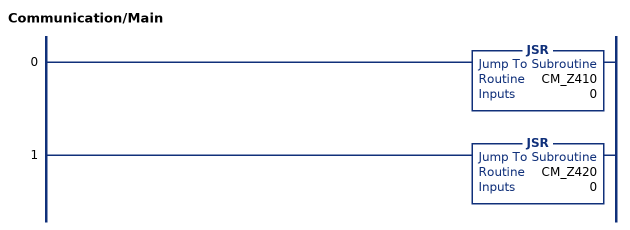
   0: JSR(CM_Z410,0);
   1: JSR(CM_Z420,0);
END_ROUTINE
END_PROGRAM

PROGRAM Initialize   (* main routine Main *)
VAR
   CapsConveyor_INIT : UDT_CapsConveyor_ZC[10]; {access None}
   Conveyor_INIT : UDT_StandConv[29]; {access None}
   M302SpeedUp_INIT : MAC_SpeedUp := (tmON_TimeControlSnap[0].PRE := 30000, tmON_TimeControlSnap[1].PRE := 30000); {constant, access None}
   M307ASpeedUp_INIT : MAC_SpeedUp := (tmON_TimeControlSnap[0].PRE := 30000, tmON_TimeControlSnap[1].PRE := 30000); {constant, access None}
   M30xTrimDeck_INIT : MAC_TrimmingDeck; {constant}
   M30xTrimWheels_INIT : MAC_TrimmingWheels[4]; {constant, access None}
        [1]   // M303 DW
        [2]   // M304 UP
        [3]   // M304 DW
        [0]   // M303 UP
   M310Popup_INIT : MAC_Popup_ZC[2]; {constant, access None}
        [0].PH_x.24   // Unload to stacker
        [0].PH_x.0   // Lift
        [0].PH_x.27   // End load to stacker
        [0].PH_x.16   // Squaring
        [0].PH_x.11   // Unload on side leg to opposite operator side
        [0].PH_x.15   // End unload to side leg
        [0].PH_x.19   // Positiong after squaring
        [0].PH_x.28   // Load from stacker
        [0].PH_x.3   // End lift
        [0].PH_x.31   // End load from stacker
        [0].PH_x.4   // Descent
        [0].PH_x.7   // End descent
        [0].PH_x.8   // Unload on side leg to operator side
        [1].PH_x.0   // Lift
        [1].PH_x.11   // Unload on side leg to opposite operator side
        [1].PH_x.15   // End unload to side leg
        [1].PH_x.16   // Squaring
        [1].PH_x.19   // Positiong after squaring
        [1].PH_x.24   // Unload to stacker
        [1].PH_x.27   // End load to stacker
        [1].PH_x.28   // Load from stacker
        [1].PH_x.3   // End lift
        [1].PH_x.31   // End load from stacker
        [1].PH_x.4   // Descent
        [1].PH_x.7   // End descent
        [1].PH_x.8   // Unload on side leg to operator side
   M315Popup_INIT : MAC_Popup_ZC[2]; {constant, access None}
        [0].PH_x.0   // Lift
        [0].PH_x.11   // Unload on side leg to opposite operator side
        [0].PH_x.15   // End unload to side leg
        [0].PH_x.16   // Squaring
        [0].PH_x.19   // Positiong after squaring
        [0].PH_x.24   // Unload to stacker
        [0].PH_x.27   // End load to stacker
        [0].PH_x.28   // Load from stacker
        [0].PH_x.3   // End lift
        [0].PH_x.31   // End load from stacker
        [0].PH_x.4   // Descent
        [0].PH_x.7   // End descent
        [0].PH_x.8   // Unload on side leg to operator side
        [1].PH_x.0   // Lift
        [1].PH_x.11   // Unload on side leg to opposite operator side
        [1].PH_x.15   // End unload to side leg
        [1].PH_x.16   // Squaring
        [1].PH_x.19   // Positiong after squaring
        [1].PH_x.24   // Unload to stacker
        [1].PH_x.27   // End load to stacker
        [1].PH_x.28   // Load from stacker
        [1].PH_x.3   // End lift
        [1].PH_x.31   // End load from stacker
        [1].PH_x.4   // Descent
        [1].PH_x.7   // End descent
        [1].PH_x.8   // Unload on side leg to operator side
   M350Popup_INIT : MAC_Popup_ZC; {access Read Only}
   Tracking_INIT : UDT_Tracking; {access None}
   Z301_INIT : MAC_Zone_ML := (tmON_ResetAlarm.PRE := 2000, tmON_24Vdc.PRE := 2000, tmON_400Vca.PRE := 2000, tmON_EmergencyOK.PRE := 2000, tmON_Cycle.PRE := 15000, tmON_ForceStop.PRE := 2000, tmON_AllowStopCleaning.PRE := 2000, tmON_CycleAcousticAlarm.PRE := 15000, tmON_ConveyorsNotOK.PRE := 2000, tmON_StopCycleForFaults.PRE := 2000, tmON_StopCycleForSaturation.PRE := 2000); {constant, access None}
END_VAR

ROUTINE Main   (* ladder *)
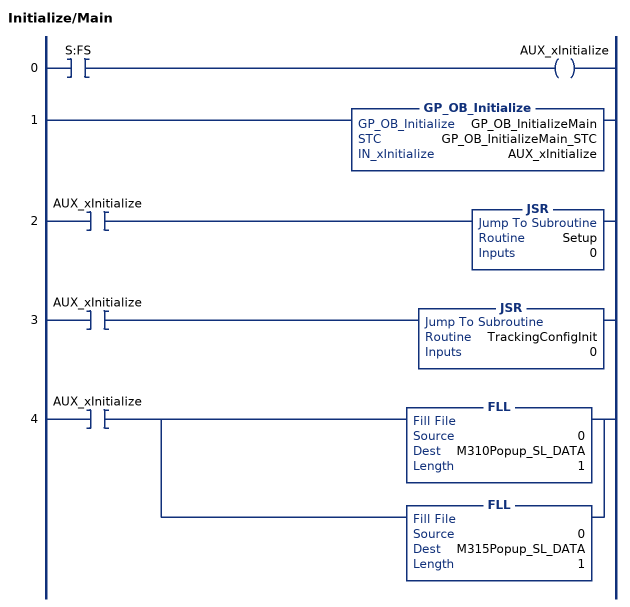
   0: XIC(S:FS)OTE(AUX_xInitialize);
   1: GP_OB_Initialize(GP_OB_InitializeMain,GP_OB_InitializeMain_STC,AUX_xInitialize);
   2: XIC(AUX_xInitialize)JSR(Setup,0);
   3: XIC(AUX_xInitialize)JSR(TrackingConfigInit,0);
   4: XIC(AUX_xInitialize)[FLL(0,M310Popup_SL_DATA,1) ,FLL(0,M315Popup_SL_DATA,1) ];
END_ROUTINE

ROUTINE Setup   (* structured text *)
   //Upload initialize parameters
   //Main line
   (*COP(Z301,Z301_INIT,1);
   COP(Z302,Z302_INIT,1);
   COP(Z303,Z303_INIT,1);
   COP(M301SpeedUp,M301SpeedUp_INIT,1);
   COP(M313SpeedUp,M313SpeedUp_INIT,1);
   COP(M31xConveyor[0],M31xConveyor_INIT[0],CONST_tPlant.dZ1ConveyorNumber);
   COP(M32xConveyor[0],M32xConveyor_INIT[0],CONST_tPlant.dZ2ConveyorNumber);
   COP(M33xConveyor[0],M33xConveyor_INIT[0],CONST_tPlant.dZ3ConveyorNumber);
   COP(M303TrimDeck,M303TrimDeck_INIT,1);
   COP(M303xTrimWheel[0],M303xTrimWheel_INIT[0],CONST_tPlant.dTrimWheelsNumber);
   COP(M311ASplitBar,M311ASplitBar_INIT,1);
   COP(M311BSeparatorRolls,M311BSeparatorRolls_INIT,1);
   COP(M385PowderMachine,M385_INIT,1);
   COP(M314AInputBreaker,M314AInputBreaker_INIT,1);
   COP(M320AInputBreaker,M320AInputBreaker_INIT,1);
   COP(M317Popup[0],M317Popup_INIT[0],2);
   COP(M325Popup[0],M325Popup_INIT[0],2);
   COP(M323Popup,M323Popup_INIT,1);
   COP(M327Popup,M327Popup_INIT,1);
   COP(M314BBreaker,M314BBreaker_INIT,1);
   COP(M320BBreaker,M320BBreaker_INIT,1);
   COP(M390Breaker,M390Breaker_INIT,1);*)
   
   //Download initialize parameters
   //Main line
   //COP(M31xConveyor_INIT[0],M31xConveyor[0],CONST_tPlant.dZ1ConveyorNumber);
   //COP(M32xConveyor_INIT[0],M32xConveyor[0],CONST_tPlant.dZ2ConveyorNumber);
   //COP(M33xConveyor_INIT[0],M33xConveyor[0],CONST_tPlant.dZ3ConveyorNumber);
   COP(Conveyor_INIT[0],Z300_Conveyor[0],CONST_tPlant.dNumOfConveyors);
   FOR TMP_dIndexConv := 0 TO CONST_tPlant.dNumOfConveyors - 1 DO
   	FOR TMP_dIndexCapConv := 0 TO CONST_tPlant.dNumCapsConveyor - 1 DO
   		COP(AUX_tCapsConveyor_NULL,Z300_LineTracking.rgtTrkConv[TMP_dIndexConv].Cap[TMP_dIndexCapConv],1);
   	END_FOR;
   END_FOR;
   COP(Z301_INIT,Z301,1);
   Z301.ST_xSelAutoMode:=1;
   
   COP(M302SpeedUp_INIT,M302SpeedUp,1);
   COP(M307ASpeedUp_INIT,M307ASpeedUp,1);
   FOR TMP_dIndex := 0 TO CONST_tPlant.dTrimDeckNumber - 1 DO
   	COP(M30xTrimDeck_INIT,M30xTrimDeck[TMP_dIndex],1);
   END_FOR;
   FOR TMP_dIndex := 0 TO CONST_tPlant.dTrimWheelsNumber - 1 DO
   	COP(M30xTrimWheels_INIT[0],M30xTrimWheel[TMP_dIndex],1);
   END_FOR;
   
   COP(M350Popup_INIT,M350Popup,1);
   
   FOR TMP_dIndex := 0 TO 1 DO
   	COP(M310Popup_INIT[0],M310Popup[TMP_dIndex],1);
   	COP(M315Popup_INIT[0],M315Popup[TMP_dIndex],1);
   END_FOR;
   
   (*//Preset time on indexed machines
   //Load preset time on M31xConveyors
   FOR TMP_dPnt1:=0 TO CONST_tPlant.dZ1ConveyorNumber - 1 DO
   	M31xConveyor[TMP_dPnt1].tmON_Wait.PRE:=0;
   	M31xConveyor[TMP_dPnt1].tmON_SyncTimeout.PRE:=20000;
   	M31xConveyor[TMP_dPnt1].tmOF_SyncTimeout.PRE:=2000;
   	M31xConveyor[TMP_dPnt1].tmON_PhFilter.PRE:=200;
   	IF M31xConveyor[TMP_dPnt1].CONST_dMotorNumber > 0 THEN
   		TMP_d:=M31xConveyor[TMP_dPnt1].CONST_dMotorNumber;
   	ELSE
   		TMP_d:=1;
   	END_IF;
   	FOR TMP_dPnt2:=0 TO TMP_d - 1 DO
   		M31xConveyor[TMP_dPnt1].tmON_FeedbackTimeOut[TMP_dPnt2].PRE:=1500;
   		M31xConveyor[TMP_dPnt1].tmOF_DriveEnable[TMP_dPnt2].PRE:=20000;
   	END_FOR;
   END_FOR;
   
   //Load preset time on M32xConveyors
   FOR TMP_dPnt1:=0 TO CONST_tPlant.dZ2ConveyorNumber - 1 DO
   	M32xConveyor[TMP_dPnt1].tmON_Wait.PRE:=0;
   	M32xConveyor[TMP_dPnt1].tmON_SyncTimeout.PRE:=20000;
   	M32xConveyor[TMP_dPnt1].tmOF_SyncTimeout.PRE:=2000;
   	M32xConveyor[TMP_dPnt1].tmON_PhFilter.PRE:=200;
   	IF M32xConveyor[TMP_dPnt1].CONST_dMotorNumber > 0 THEN
   		TMP_d:=M32xConveyor[TMP_dPnt1].CONST_dMotorNumber;
   	ELSE
   		TMP_d:=1;
   	END_IF;
   	FOR TMP_dPnt2:=0 TO TMP_d - 1 DO
   		M32xConveyor[TMP_dPnt1].tmON_FeedbackTimeOut[TMP_dPnt2].PRE:=1500;
   		M32xConveyor[TMP_dPnt1].tmOF_DriveEnable[TMP_dPnt2].PRE:=20000;
   	END_FOR;
   END_FOR;
   
   //Load preset time on M33xConveyors
   FOR TMP_dPnt1:=0 TO CONST_tPlant.dZ2ConveyorNumber - 1 DO
   	M33xConveyor[TMP_dPnt1].tmON_Wait.PRE:=0;
   	M33xConveyor[TMP_dPnt1].tmON_SyncTimeout.PRE:=20000;
   	M33xConveyor[TMP_dPnt1].tmOF_SyncTimeout.PRE:=2000;
   	M33xConveyor[TMP_dPnt1].tmON_PhFilter.PRE:=200;
   	IF M33xConveyor[TMP_dPnt1].CONST_dMotorNumber > 0 THEN
   		TMP_d:=M33xConveyor[TMP_dPnt1].CONST_dMotorNumber;
   	ELSE
   		TMP_d:=1;
   	END_IF;
   	FOR TMP_dPnt2:=0 TO TMP_d - 1 DO
   		M33xConveyor[TMP_dPnt1].tmON_FeedbackTimeOut[TMP_dPnt2].PRE:=1500;
   		M33xConveyor[TMP_dPnt1].tmOF_DriveEnable[TMP_dPnt2].PRE:=20000;
   	END_FOR;
   END_FOR;*)
   
   //Load preset time on M30xTrimDeck
   FOR TMP_d :=0 TO CONST_tPlant.dTrimDeckNumber - 1 DO
   	M30xTrimDeck[TMP_d].tmON_EncPreset[0].PRE:=3000;
   	M30xTrimDeck[TMP_d].tmON_EncPreset[1].PRE:=3000;
   	M30xTrimDeck[TMP_d].tmON_CheckEncoderTimeOut[0].PRE:=1000;
   	M30xTrimDeck[TMP_d].tmON_CheckEncoderTimeOut[1].PRE:=1000;
   	M30xTrimDeck[TMP_d].tmON_FeedbackTimeOut[0].PRE:=2500;
   	M30xTrimDeck[TMP_d].tmON_FeedbackTimeOut[1].PRE:=2500;
   	M30xTrimDeck[TMP_d].tmOF_DriveEnable[0].PRE:=30000;
   	M30xTrimDeck[TMP_d].tmOF_DriveEnable[1].PRE:=30000;
   	M30xTrimDeck[TMP_d].tmOF_DelayOnChangeDirection[0].PRE:=500;
   	M30xTrimDeck[TMP_d].tmOF_DelayOnChangeDirection[1].PRE:=500;
   	M30xTrimDeck[TMP_d].tmOF_DelayOnChangeDirection[2].PRE:=500;
   	M30xTrimDeck[TMP_d].tmOF_DelayOnChangeDirection[3].PRE:=500;
   	M30xTrimDeck[TMP_d].tmON_Wait.PRE:=0;
   END_FOR;
   
   //Load preset time on M30xTrimWheels
   FOR TMP_d :=0 TO CONST_tPlant.dTrimWheelsNumber - 1 DO
   	M30xTrimWheel[TMP_d].tmON_TrimWheelTimeOut[0].PRE:=2500;
   	M30xTrimWheel[TMP_d].tmON_TrimWheelTimeOut[1].PRE:=2500;
   	M30xTrimWheel[TMP_d].tmON_Wait[0].PRE:=0;
   	M30xTrimWheel[TMP_d].tmON_Wait[1].PRE:=0;
   END_FOR;
   
   //Load preset time M317Popup
   M310Popup[0].tmON_LiftingTimeOut.PRE := 2000;
   M310Popup[0].tmON_LiftingFeedbackTimeOut.PRE := 1000;
   M310Popup[0].tmOF_WaitBothEndLift.PRE := 1500;
   M310Popup[0].tmON_ReentryPlate.PRE := 200;
   M310Popup[0].tmON_Positioning.PRE := 40;
   M310Popup[1].tmON_LiftingTimeOut.PRE := 2000;
   M310Popup[1].tmON_LiftingFeedbackTimeOut.PRE := 1000;
   M310Popup[1].tmOF_WaitBothEndLift.PRE := 1500;
   M310Popup[1].tmON_ReentryPlate.PRE := 200;
   M310Popup[1].tmON_Positioning.PRE := 40;
   
   //Load preset time M325Popup
   M315Popup[0].tmON_LiftingTimeOut.PRE := 2000;
   M315Popup[0].tmON_LiftingFeedbackTimeOut.PRE := 1000;
   M315Popup[0].tmOF_WaitBothEndLift.PRE := 1500;
   M315Popup[0].tmON_ReentryPlate.PRE := 200;
   M315Popup[0].tmON_Positioning.PRE := 40;
   M315Popup[1].tmON_LiftingTimeOut.PRE := 2000;
   M315Popup[1].tmON_LiftingFeedbackTimeOut.PRE := 1000;
   M315Popup[1].tmOF_WaitBothEndLift.PRE := 1500;
   M315Popup[1].tmON_ReentryPlate.PRE := 200;
   M315Popup[1].tmON_Positioning.PRE := 40;
   
END_ROUTINE

ROUTINE TrackingConfigInit   (* structured text *)
   
   Z300_dStartTrackingPosition := 0;
   Z300_LineTracking.rgtTrkConv[0].dStartPosition_cmm := Z300_dStartTrackingPosition;
   Z300_LineTracking.rgtTrkConv[0].dEndPosition_cmm := Z300_dStartTrackingPosition + Z300_Conveyor_Conf[0].dLengthConveyor_cmm;
   size(Z300_LineTracking.rgtTrkConv[0],0,TMP_dLineSize);
   FOR TMP_dIndexConv := 1 TO TMP_dLineSize - 1 DO
   	Z300_LineTracking.rgtTrkConv[TMP_dIndexConv].dStartPosition_cmm := Z300_LineTracking.rgtTrkConv[TMP_dIndexConv - 1].dEndPosition_cmm;
   	Z300_LineTracking.rgtTrkConv[TMP_dIndexConv].dEndPosition_cmm := Z300_LineTracking.rgtTrkConv[TMP_dIndexConv].dStartPosition_cmm + Z300_Conveyor_Conf[TMP_dIndexConv].dLengthConveyor_cmm;
   END_FOR;
   Z300_dEndTrackingPosition := Z300_LineTracking.rgtTrkConv[TMP_dLineSize - 1].dEndPosition_cmm;
   
END_ROUTINE
END_PROGRAM

PROGRAM MainProgram   (* main routine MainRoutine *)

ROUTINE _10_MCP_I   (* ladder *)
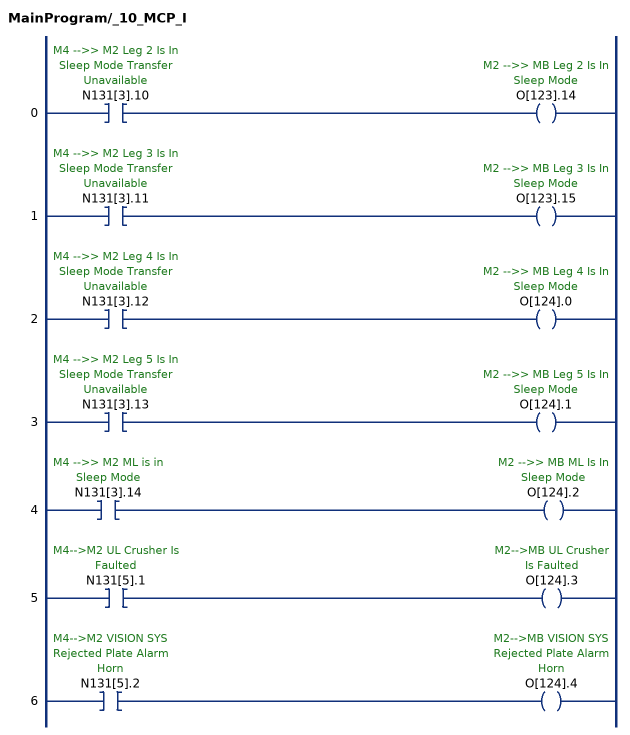
   0: XIC(N131[3].10)OTE(O[123].14);
   1: XIC(N131[3].11)OTE(O[123].15);
   2: XIC(N131[3].12)OTE(O[124].0);
   3: XIC(N131[3].13)OTE(O[124].1);
   4: XIC(N131[3].14)OTE(O[124].2);
   5: XIC(N131[5].1)OTE(O[124].3);
   6: XIC(N131[5].2)OTE(O[124].4);
END_ROUTINE

ROUTINE _12_MCP_K   (* ladder *)
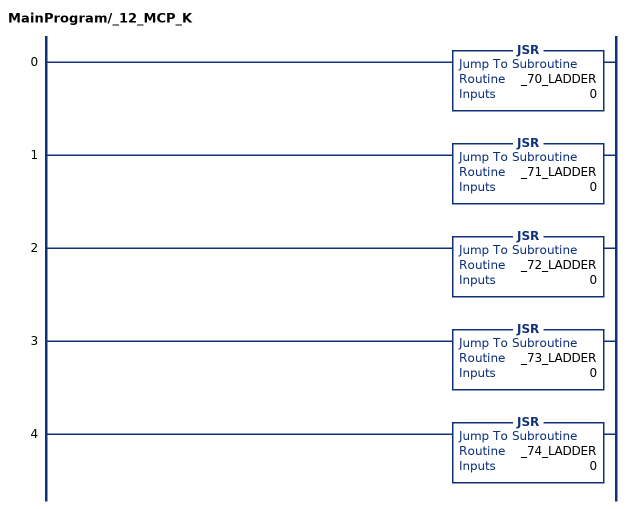
   0: JSR(_70_LADDER,0);
   1: JSR(_71_LADDER,0);
   2: JSR(_72_LADDER,0);
   3: JSR(_73_LADDER,0);
   4: JSR(_74_LADDER,0);
END_ROUTINE

ROUTINE _26_ADAPTER   (* ladder *)
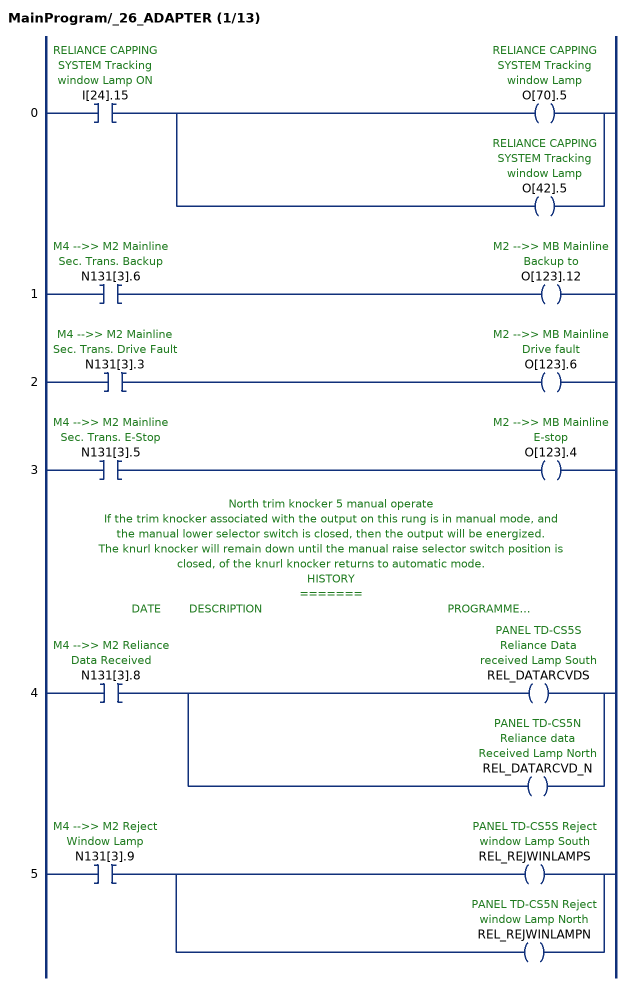
   0: XIC(I[24].15)[OTE(O[70].5) ,OTE(O[42].5) ];
   1: XIC(N131[3].6)OTE(O[123].12);
   2: XIC(N131[3].3)OTE(O[123].6);
   3: XIC(N131[3].5)OTE(O[123].4);
   // North trim knocker 5 manual operate
   // If the trim knocker associated with the output on this rung is in manual mode, and
   // the manual lower selector switch is closed, then the output will be energized.
   // The knurl knocker will remain down until the manual raise selector switch position is
   // closed, of the knurl knocker returns to automatic mode.
   // HISTORY
   // =======
   // DATE        DESCRIPTION                                                     PROGRAMMER
   // ====        ===========                                                     ==========
   // 2/29/96     Entered rung as designed                                        WAS
   // 3/1/96      Added these comments                                            WAS
   4: XIC(N131[3].8)[OTE(REL_DATARCVDS) ,OTE(REL_DATARCVD_N) ];
   5: XIC(N131[3].9)[OTE(REL_REJWINLAMPS) ,OTE(REL_REJWINLAMPN) ];
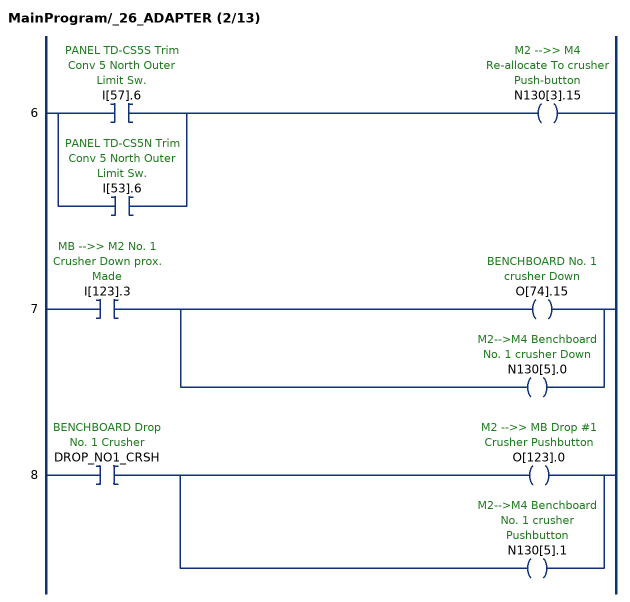
   6: [XIC(I[57].6) ,XIC(I[53].6) ]OTE(N130[3].15);
   7: XIC(I[123].3)[OTE(O[74].15) ,OTE(N130[5].0) ];
   8: XIC(DROP_NO1_CRSH)[OTE(O[123].0) ,OTE(N130[5].1) ];
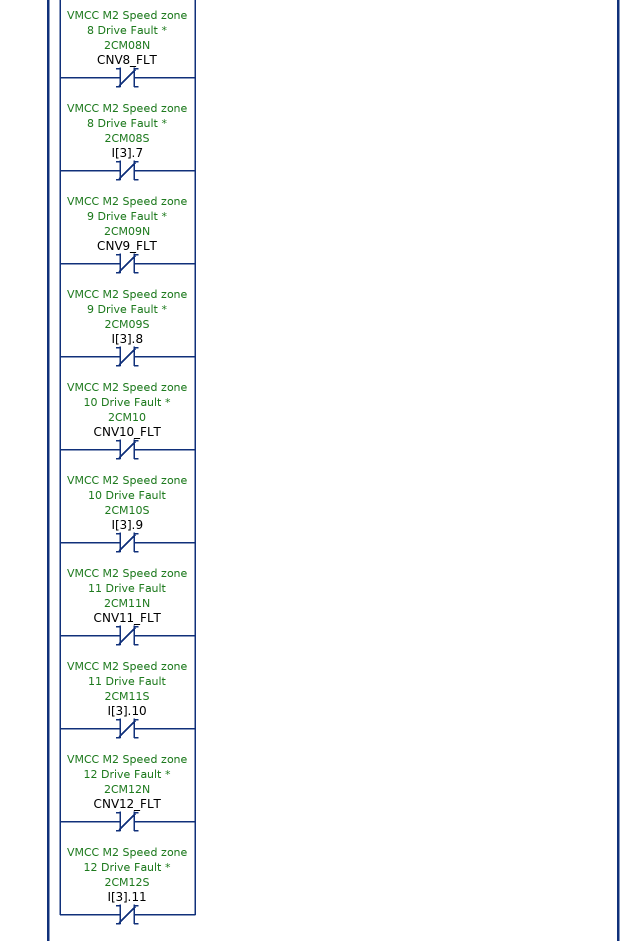
   9: [XIO(CNV1_FLT) ,XIO(CNV2_FLT) ,XIO(CNV3_FLT) ,XIO(CNV4_FLT) ,XIO(I[3].3) ,XIO(CNV5_FLT) ,XIO(I[3].4) ,XIO(CNV6_FLT) ,XIO(I[3].5) ,XIO(CNV7_FLT) ,XIO(I[3].6) ,XIO(CNV8_FLT) ,XIO(I[3].7) ,XIO(CNV9_FLT) ,XIO(I[3].8) ,XIO(CNV10_FLT) ,XIO(I[3].9) ,XIO(CNV11_FLT) ,XIO(I[3].10) ,XIO(CNV12_FLT) ,XIO(I[3].11) ]TON(T4[33],?,?);
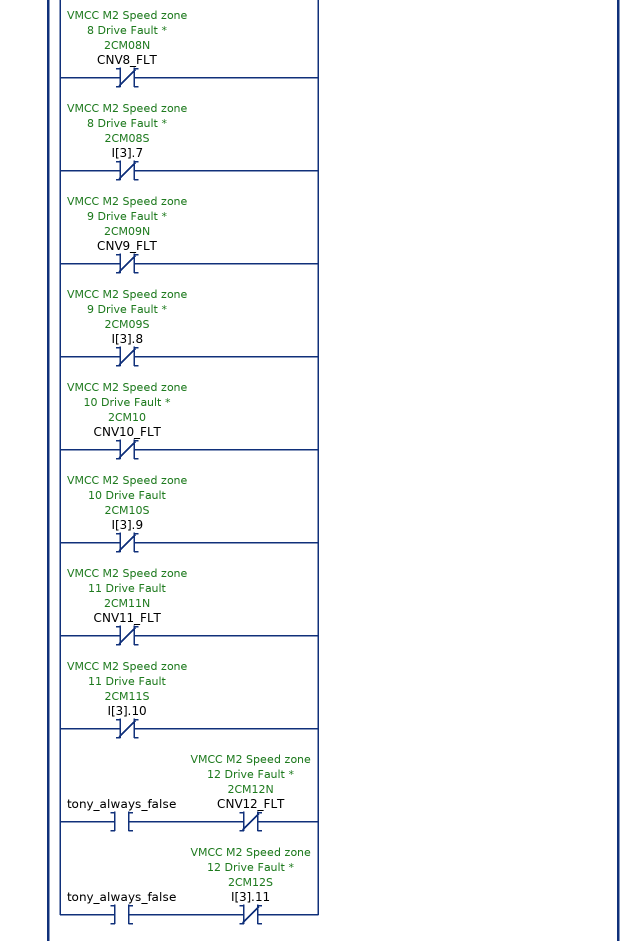
   10: [XIO(CNV1_FLT) ,XIO(CNV2_FLT) ,XIO(CNV3_FLT) ,XIO(CNV4_FLT) ,XIO(I[3].3) ,XIO(CNV5_FLT) ,XIO(I[3].4) ,XIO(CNV6_FLT) ,XIO(I[3].5) ,XIO(CNV7_FLT) ,XIO(I[3].6) ,XIO(CNV8_FLT) ,XIO(I[3].7) ,XIO(CNV9_FLT) ,XIO(I[3].8) ,XIO(CNV10_FLT) ,XIO(I[3].9) ,XIO(CNV11_FLT) ,XIO(I[3].10) ,XIC(tony_always_false) XIO(CNV12_FLT) ,XIC(tony_always_false) XIO(I[3].11) ]TON(T4[33],?,?);
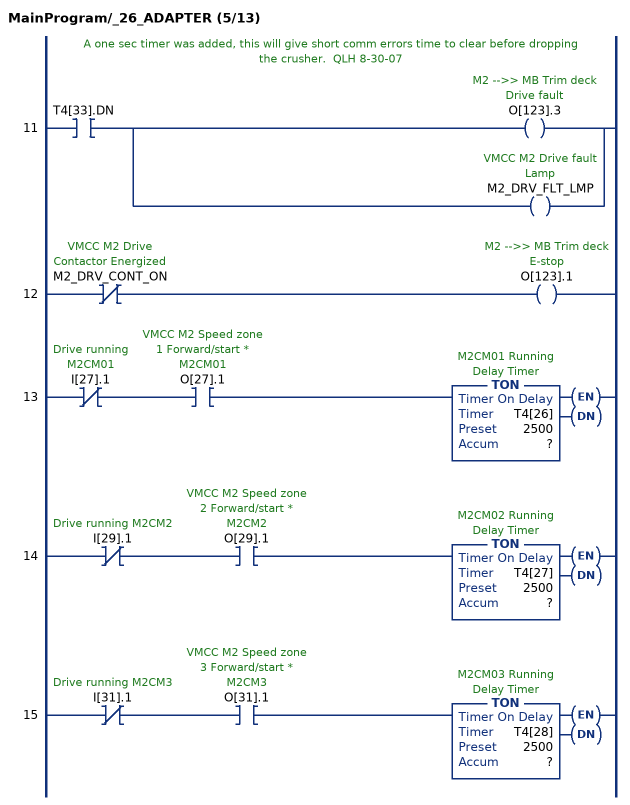
   // A one sec timer was added, this will give short comm errors time to clear before dropping the crusher.  QLH 8-30-07
   11: XIC(T4[33].DN)[OTE(O[123].3) ,OTE(M2_DRV_FLT_LMP) ];
   12: XIO(M2_DRV_CONT_ON)OTE(O[123].1);
   13: XIO(I[27].1)XIC(O[27].1)TON(T4[26],?,?);
   14: XIO(I[29].1)XIC(O[29].1)TON(T4[27],?,?);
   15: XIO(I[31].1)XIC(O[31].1)TON(T4[28],?,?);
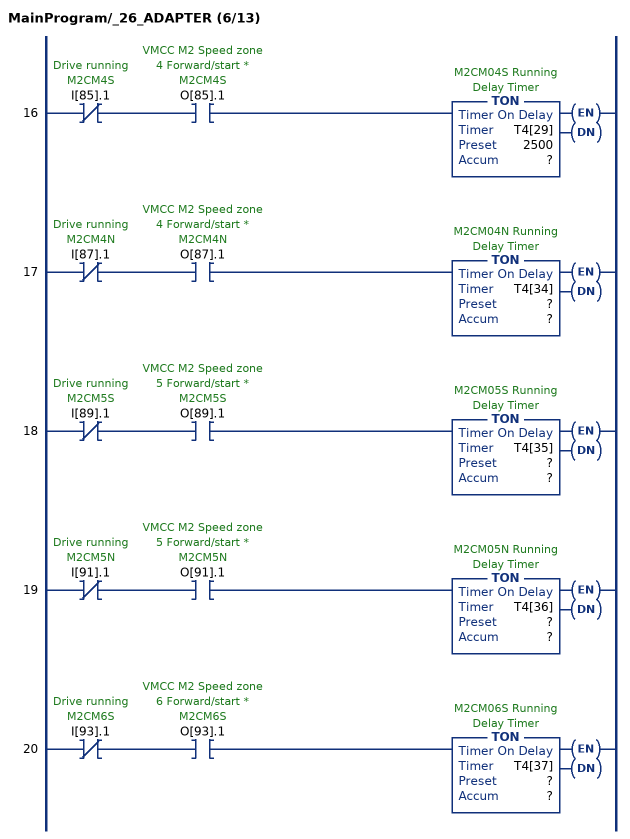
   16: XIO(I[85].1)XIC(O[85].1)TON(T4[29],?,?);
   17: XIO(I[87].1)XIC(O[87].1)TON(T4[34],?,?);
   18: XIO(I[89].1)XIC(O[89].1)TON(T4[35],?,?);
   19: XIO(I[91].1)XIC(O[91].1)TON(T4[36],?,?);
   20: XIO(I[93].1)XIC(O[93].1)TON(T4[37],?,?);
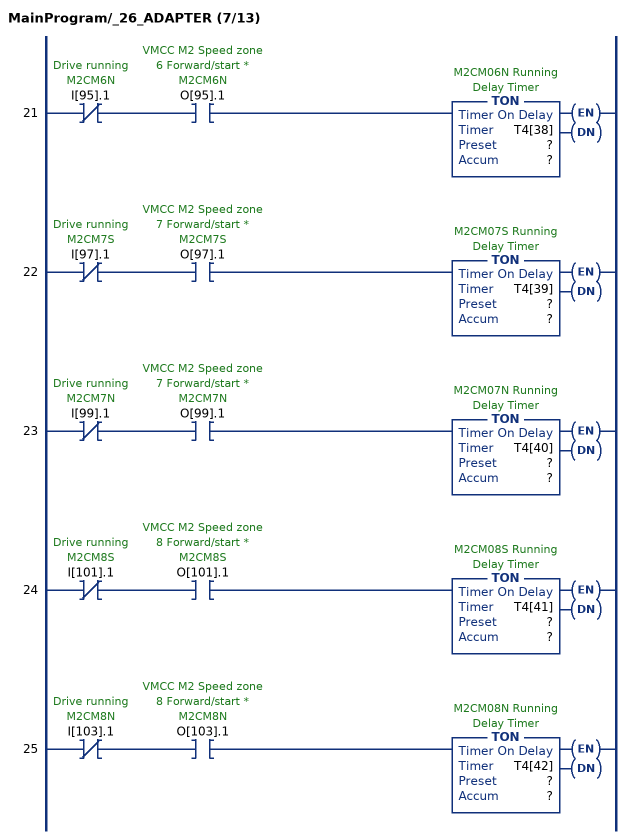
   21: XIO(I[95].1)XIC(O[95].1)TON(T4[38],?,?);
   22: XIO(I[97].1)XIC(O[97].1)TON(T4[39],?,?);
   23: XIO(I[99].1)XIC(O[99].1)TON(T4[40],?,?);
   24: XIO(I[101].1)XIC(O[101].1)TON(T4[41],?,?);
   25: XIO(I[103].1)XIC(O[103].1)TON(T4[42],?,?);
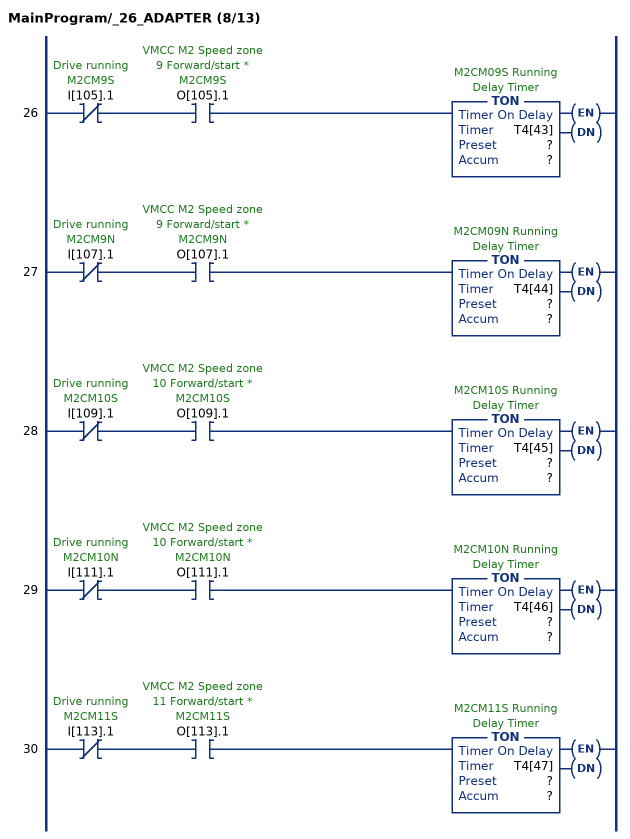
   26: XIO(I[105].1)XIC(O[105].1)TON(T4[43],?,?);
   27: XIO(I[107].1)XIC(O[107].1)TON(T4[44],?,?);
   28: XIO(I[109].1)XIC(O[109].1)TON(T4[45],?,?);
   29: XIO(I[111].1)XIC(O[111].1)TON(T4[46],?,?);
   30: XIO(I[113].1)XIC(O[113].1)TON(T4[47],?,?);
